   Group "Group" at 455,41 size 373x50
   Button "HmiScreenItemData_8" at 469,45 size 355x40; TextOn 'Back'; TextOff 'Text'
   TextField "Screen title" at 455,41 size 373x50; Text 'Screen title'

screen "BC Max Step Times" 1280x800, template "Template"
   on GenerateScreen: "TitleUpdater"()
   Button "HmiScreenItemData_1" at 1,1 size 150x43; TextOn 'Back'; TextOff 'Commissioning'
      on Release: ActivateScreen("Commissioning Main Page", 0)
   Button "Button_1" at 21,736 size 161x32; TextOff 'Back'
      on Activate: ActivateScreen("IGG Process Times", 0)
   TextField "Text field_25" at 83,285 size 286x22; Text 'Step 040'
   TextField "Text field_29" at 383,118 size 77x20; Text 'Time (ms)'
   TextField "Text field_33" at 83,312 size 286x22; Text 'Step 050'
   IOField "I/O field_58" at 382,312 size 60x22; Authorization "Parameter Change"; FormatPattern s9999999999
      ProcessValue <- "86_Times_STEP_MAX_TIME_STP_050(1)"
   TextField "Text field_35" at 83,367 size 286x22; Text 'Step 070'
   TextField "Text field_65" at 83,144 size 286x22; Text 'Step 001'
   TextField "Text field_67" at 83,173 size 286x22; Text 'Step 005'
   TextField "Text field_69" at 83,200 size 286x22; Text 'Step 010'
   TextField "Text field_71" at 83,229 size 286x22; Text 'Step 020'
   TextField "Text field_73" at 83,257 size 286x22; Text 'Step 030'
   TextField "Text field_42" at 83,118 size 89x20; Text 'Description'
   IOField "I/O field_128" at 382,144 size 60x22; Authorization "Parameter Change"; FormatPattern s9999999999
      ProcessValue <- "86_Times_STEP_MAX_TIME_STP_001(1)"
   IOField "I/O field_133" at 382,173 size 60x22; Authorization "Parameter Change"; FormatPattern s9999999999
      ProcessValue <- "86_Times_STEP_MAX_TIME_STP_005(1)"
   IOField "I/O field_138" at 382,200 size 60x22; Authorization "Parameter Change"; FormatPattern s9999999999
      ProcessValue <- "86_Times_STEP_MAX_TIME_STP_010(1)"
   IOField "I/O field_148" at 382,257 size 60x22; Authorization "Parameter Change"; FormatPattern s9999999999
      ProcessValue <- "86_Times_STEP_MAX_TIME_STP_030(1)"
   IOField "I/O field_64" at 382,367 size 60x22; Authorization "Parameter Change"; FormatPattern s9999999999
      ProcessValue <- "86_Times_STEP_MAX_TIME_STP_070(1)"
   TextField "Text field_53" at 82,92 size 247x26; Text 'BC Maximum Step Times'
   IOField "I/O field_5" at 382,229 size 60x22; Authorization "Parameter Change"; FormatPattern s9999999999
      ProcessValue <- "86_Times_STEP_MAX_TIME_STP_020(1)"
   TextField "Text field_1" at 83,340 size 286x22; Text 'Step 060'
   IOField "I/O field_2" at 382,340 size 60x22; Authorization "Parameter Change"; FormatPattern s9999999999
      ProcessValue <- "86_Times_STEP_MAX_TIME_STP_060(1)"
   TextField "Text field_2" at 461,286 size 286x22; Text 'Step 240'
   TextField "Text field_3" at 750,119 size 77x20; Text 'Time (ms)'
   TextField "Text field_4" at 461,313 size 286x22; Text 'Step 250'
   IOField "I/O field_1" at 758,312 size 60x22; Authorization "Parameter Change"; FormatPattern s9999999999
      ProcessValue <- "86_Times_STEP_MAX_TIME_STP_250(1)"
   TextField "Text field_5" at 461,368 size 286x22; Text 'Step 270'
   TextField "Text field_6" at 461,145 size 286x22; Text 'Step 190'
   TextField "Text field_7" at 461,174 size 286x22; Text 'Step 200'
   TextField "Text field_8" at 461,201 size 286x22; Text 'Step 210'
   TextField "Text field_9" at 461,230 size 286x22; Text 'Step 220'
   TextField "Text field_10" at 461,258 size 286x22; Text 'Step 230'
   TextField "Text field_11" at 461,119 size 89x20; Text 'Description'
   IOField "I/O field_3" at 758,145 size 60x22; Authorization "Parameter Change"; FormatPattern s9999999999
      ProcessValue <- "86_Times_STEP_MAX_TIME_STP_190(1)"
   IOField "I/O field_4" at 758,174 size 60x22; Authorization "Parameter Change"; FormatPattern s9999999999
      ProcessValue <- "86_Times_STEP_MAX_TIME_STP_200(1)"
   IOField "I/O field_6" at 758,201 size 60x22; Authorization "Parameter Change"; FormatPattern s9999999999
      ProcessValue <- "86_Times_STEP_MAX_TIME_STP_210(1)"
   IOField "I/O field_8" at 758,258 size 60x22; Authorization "Parameter Change"; FormatPattern s9999999999
      ProcessValue <- "86_Times_STEP_MAX_TIME_STP_230(1)"
   IOField "I/O field_9" at 758,367 size 60x22; Authorization "Parameter Change"; FormatPattern s9999999999
      ProcessValue <- "86_Times_STEP_MAX_TIME_STP_270(1)"
   IOField "I/O field_10" at 758,230 size 60x22; Authorization "Parameter Change"; FormatPattern s9999999999
      ProcessValue <- "86_Times_STEP_MAX_TIME_STP_220(1)"
   TextField "Text field_13" at 461,341 size 286x22; Text 'Step 260'
   IOField "I/O field_11" at 758,340 size 60x22; Authorization "Parameter Change"; FormatPattern s9999999999
      ProcessValue <- "86_Times_STEP_MAX_TIME_STP_260(1)"
   TextField "Text field_14" at 83,398 size 286x22; Text 'Step 080'
   IOField "I/O field_12" at 382,398 size 60x22; Authorization "Parameter Change"; FormatPattern s9999999999
      ProcessValue <- "86_Times_STEP_MAX_TIME_STP_080(1)"
   TextField "Text field_15" at 83,426 size 286x22; Text 'Step 090'
   IOField "I/O field_13" at 382,426 size 60x22; Authorization "Parameter Change"; FormatPattern s9999999999
      ProcessValue <- "86_Times_STEP_MAX_TIME_STP_090(1)"
   TextField "Text field_16" at 83,453 size 286x22; Text 'Step 100'
   IOField "I/O field_14" at 382,453 size 60x22; Authorization "Parameter Change"; FormatPattern s9999999999
      ProcessValue <- "86_Times_STEP_MAX_TIME_STP_100(1)"
   IOField "I/O field_15" at 382,285 size 60x22; Authorization "Parameter Change"; FormatPattern s9999999999
      ProcessValue <- "86_Times_STEP_MAX_TIME_STP_040(1)"
   TextField "Text field_17" at 461,395 size 286x22; Text 'Step 280'
   IOField "I/O field_16" at 758,394 size 60x22; Authorization "Parameter Change"; FormatPattern s9999999999
      ProcessValue <- "86_Times_STEP_MAX_TIME_STP_280(1)"
   TextField "Text field_18" at 461,426 size 286x22; Text 'Step 290'
   IOField "I/O field_17" at 758,425 size 60x22; Authorization "Parameter Change"; FormatPattern s9999999999
      ProcessValue <- "86_Times_STEP_MAX_TIME_STP_290(1)"
   TextField "Text field_19" at 461,453 size 286x22; Text 'Step 300'
   IOField "I/O field_18" at 758,452 size 60x22; Authorization "Parameter Change"; FormatPattern s9999999999
      ProcessValue <- "86_Times_STEP_MAX_TIME_STP_300(1)"
   TextField "Text field_20" at 461,483 size 286x22; Text 'Step 310'
   IOField "I/O field_19" at 758,482 size 60x22; Authorization "Parameter Change"; FormatPattern s9999999999
      ProcessValue <- "86_Times_STEP_MAX_TIME_STP_310(1)"
   TextField "Text field_21" at 461,510 size 286x22; Text 'Step 320'
   IOField "I/O field_20" at 758,509 size 60x22; Authorization "Parameter Change"; FormatPattern s9999999999
      ProcessValue <- "86_Times_STEP_MAX_TIME_STP_320(1)"
   TextField "Text field_22" at 835,145 size 286x22; Text 'Step 390'
   IOField "I/O field_21" at 1130,144 size 60x22; Authorization "Parameter Change"; FormatPattern s9999999999
      ProcessValue <- "86_Times_STEP_MAX_TIME_STP_390(1)"
   TextField "Text field_23" at 835,118 size 89x20; Text 'Description'
   TextField "Text field_24" at 1122,119 size 77x20; Text 'Time (ms)'
   TextField "Text field_26" at 835,173 size 286x22; Text 'Step 400'
   IOField "I/O field_22" at 1130,172 size 60x22; Authorization "Parameter Change"; FormatPattern s9999999999
      ProcessValue <- "86_Times_STEP_MAX_TIME_STP_400(1)"
   TextField "Text field_27" at 835,200 size 286x22; Text 'Step 410'
   IOField "I/O field_23" at 1130,199 size 60x22; Authorization "Parameter Change"; FormatPattern s9999999999
      ProcessValue <- "86_Times_STEP_MAX_TIME_STP_410(1)"
   TextField "Text field_28" at 835,230 size 286x22; Text 'Step 420'
   IOField "I/O field_24" at 1130,229 size 60x22; Authorization "Parameter Change"; FormatPattern s9999999999
      ProcessValue <- "86_Times_STEP_MAX_TIME_STP_420(1)"
   TextField "Text field_30" at 835,257 size 286x22; Text 'Step 430'
   IOField "I/O field_25" at 1130,256 size 60x22; Authorization "Parameter Change"; FormatPattern s9999999999
      ProcessValue <- "86_Times_STEP_MAX_TIME_STP_430(1)"
   TextField "Text field_31" at 835,285 size 286x22; Text 'Step 440'
   IOField "I/O field_26" at 1130,284 size 60x22; Authorization "Parameter Change"; FormatPattern s9999999999
      ProcessValue <- "86_Times_STEP_MAX_TIME_STP_440(1)"
   TextField "Text field_32" at 835,312 size 286x22; Text 'Step 450'
   IOField "I/O field_27" at 1130,311 size 60x22; Authorization "Parameter Change"; FormatPattern s9999999999
      ProcessValue <- "86_Times_STEP_MAX_TIME_STP_450(1)"
   TextField "Text field_34" at 835,341 size 286x22; Text 'Step 460'
   IOField "I/O field_28" at 1130,340 size 60x22; Authorization "Parameter Change"; FormatPattern s9999999999
      ProcessValue <- "86_Times_STEP_MAX_TIME_STP_460(1)"
   TextField "Text field_36" at 835,369 size 286x22; Text 'Step 470'
   IOField "I/O field_29" at 1130,368 size 60x22; Authorization "Parameter Change"; FormatPattern s9999999999
      ProcessValue <- "86_Times_STEP_MAX_TIME_STP_470(1)"
   TextField "Text field_37" at 835,395 size 286x22; Text 'Step 480'
   IOField "I/O field_30" at 1130,394 size 60x22; Authorization "Parameter Change"; FormatPattern s9999999999
      ProcessValue <- "86_Times_STEP_MAX_TIME_STP_480(1)"
   TextField "Text field_38" at 835,426 size 286x22; Text 'Step 490'
   IOField "I/O field_31" at 1130,425 size 60x22; Authorization "Parameter Change"; FormatPattern s9999999999
      ProcessValue <- "86_Times_STEP_MAX_TIME_STP_490(1)"
   TextField "Text field_39" at 835,452 size 286x22; Text 'Step 500'
   IOField "I/O field_32" at 1130,451 size 60x22; Authorization "Parameter Change"; FormatPattern s9999999999
      ProcessValue <- "86_Times_STEP_MAX_TIME_STP_500(1)"
   TextField "Text field_40" at 835,482 size 286x22; Text 'Step 510'
   IOField "I/O field_33" at 1130,481 size 60x22; Authorization "Parameter Change"; FormatPattern s9999999999
      ProcessValue <- "86_Times_STEP_MAX_TIME_STP_510(1)"
   TextField "Text field_41" at 835,510 size 286x22; Text 'Step 520'
   IOField "I/O field_34" at 1130,509 size 60x22; Authorization "Parameter Change"; FormatPattern s9999999999
      ProcessValue <- "86_Times_STEP_MAX_TIME_STP_520(1)"
   IOField "I/O field_7" at 758,285 size 60x22; Authorization "Parameter Change"; FormatPattern s9999999999
      ProcessValue <- "86_Times_STEP_MAX_TIME_STP_240(1)"
   TextField "Text field_43" at 83,483 size 286x22; Text 'Step 110'
   IOField "I/O field_35" at 382,483 size 60x22; Authorization "Parameter Change"; FormatPattern s9999999999
      ProcessValue <- "86_Times_STEP_MAX_TIME_STP_110(1)"
   TextField "Text field_44" at 83,510 size 286x22; Text 'Step 120'
   IOField "I/O field_36" at 382,510 size 60x22; Authorization "Parameter Change"; FormatPattern s9999999999
      ProcessValue <- "86_Times_STEP_MAX_TIME_STP_120(1)"
   TextField "Text field_45" at 461,538 size 286x22; Text 'Step 330'
   IOField "I/O field_37" at 758,537 size 60x22; Authorization "Parameter Change"; FormatPattern s9999999999
      ProcessValue <- "86_Times_STEP_MAX_TIME_STP_330(1)"
   TextField "Text field_46" at 835,538 size 286x22; Text 'Step 530'
   IOField "I/O field_38" at 1130,537 size 60x22; Authorization "Parameter Change"; FormatPattern s9999999999
      ProcessValue <- "86_Times_STEP_MAX_TIME_STP_530(1)"
   TextField "Text field_47" at 83,538 size 286x22; Text 'Step 130'
   IOField "I/O field_39" at 382,538 size 60x22; Authorization "Parameter Change"; FormatPattern s9999999999
      ProcessValue <- "86_Times_STEP_MAX_TIME_STP_130(1)"
   TextField "Text field_48" at 461,568 size 286x22; Text 'Step 340'
   IOField "I/O field_40" at 758,567 size 60x22; Authorization "Parameter Change"; FormatPattern s9999999999
      ProcessValue <- "86_Times_STEP_MAX_TIME_STP_340(1)"
   TextField "Text field_49" at 835,568 size 286x22; Text 'Step 540'
   IOField "I/O field_41" at 1130,567 size 60x22; Authorization "Parameter Change"; FormatPattern s9999999999
      ProcessValue <- "86_Times_STEP_MAX_TIME_STP_540(1)"
   TextField "Text field_50" at 83,568 size 286x22; Text 'Step 140'
   IOField "I/O field_42" at 382,568 size 60x22; Authorization "Parameter Change"; FormatPattern s9999999999
      ProcessValue <- "86_Times_STEP_MAX_TIME_STP_140(1)"
   TextField "Text field_51" at 461,599 size 286x22; Text 'Step 350'
   IOField "I/O field_43" at 758,598 size 60x22; Authorization "Parameter Change"; FormatPattern s9999999999
      ProcessValue <- "86_Times_STEP_MAX_TIME_STP_350(1)"
   TextField "Text field_52" at 835,599 size 286x22; Text 'Step 550'
   IOField "I/O field_44" at 1130,598 size 60x22; Authorization "Parameter Change"; FormatPattern s9999999999
      ProcessValue <- "86_Times_STEP_MAX_TIME_STP_550(1)"
   TextField "Text field_54" at 83,599 size 286x22; Text 'Step 150'
   IOField "I/O field_45" at 382,599 size 60x22; Authorization "Parameter Change"; FormatPattern s9999999999
      ProcessValue <- "86_Times_STEP_MAX_TIME_STP_150(1)"
   TextField "Text field_55" at 461,628 size 286x22; Text 'Step 360'
   IOField "I/O field_46" at 758,627 size 60x22; Authorization "Parameter Change"; FormatPattern s9999999999
      ProcessValue <- "86_Times_STEP_MAX_TIME_STP_360(1)"
   TextField "Text field_56" at 835,628 size 286x22; Text 'Step 560'
   IOField "I/O field_47" at 1130,627 size 60x22; Authorization "Parameter Change"; FormatPattern s9999999999
      ProcessValue <- "86_Times_STEP_MAX_TIME_STP_560(1)"
   TextField "Text field_57" at 83,628 size 286x22; Text 'Step 160'
   IOField "I/O field_48" at 382,628 size 60x22; Authorization "Parameter Change"; FormatPattern s9999999999
      ProcessValue <- "86_Times_STEP_MAX_TIME_STP_160(1)"
   TextField "Text field_58" at 461,657 size 286x22; Text 'Step 370'
   IOField "I/O field_49" at 758,656 size 60x22; Authorization "Parameter Change"; FormatPattern s9999999999
      ProcessValue <- "86_Times_STEP_MAX_TIME_STP_370(1)"
   TextField "Text field_59" at 835,657 size 286x22; Text 'Step 570'
   IOField "I/O field_50" at 1130,656 size 60x22; Authorization "Parameter Change"; FormatPattern s9999999999
      ProcessValue <- "86_Times_STEP_MAX_TIME_STP_570(1)"
   TextField "Text field_60" at 83,657 size 286x22; Text 'Step 170'
   IOField "I/O field_51" at 382,657 size 60x22; Authorization "Parameter Change"; FormatPattern s9999999999
      ProcessValue <- "86_Times_STEP_MAX_TIME_STP_170(1)"
   TextField "Text field_61" at 461,687 size 286x22; Text 'Step 380'
   IOField "I/O field_52" at 758,686 size 60x22; Authorization "Parameter Change"; FormatPattern s9999999999
      ProcessValue <- "86_Times_STEP_MAX_TIME_STP_380(1)"
   TextField "Text field_63" at 83,687 size 286x22; Text 'Step 180'
   IOField "I/O field_54" at 382,687 size 60x22; Authorization "Parameter Change"; FormatPattern s9999999999
      ProcessValue <- "86_Times_STEP_MAX_TIME_STP_180(1)"
   Group "Group" at 455,41 size 373x50
   Button "HmiScreenItemData_8" at 469,45 size 355x40; TextOn 'Back'; TextOff 'Text'
   TextField "Screen title" at 455,41 size 373x50; Text 'Screen title'

screen "05 Alarm Buffer" 1280x800, template "Template"
   AlarmView "Alarm view_1" at 8,61 size 1258x729
   Button "HmiScreenItemData_2" at 143,2 size 139x43; TextOn 'Back'; TextOff 'Alarm'
      on Release: ActivateScreen("04 Alarm Log", 0)
   Button "HmiScreenItemData_5" at 1,2 size 139x43; TextOn 'Back'; TextOff 'Main Index'
      on Release: ActivateScreen("02 Main Index", 0)
   Button "HmiScreenItemData_4" at 1138,1 size 139x43; TextOn 'I&A Compressor Ok'; TextOff 'Back'
      on Release: function_efd93a16()

screen "08 BTCS MAIN" 1280x800, template "Template"
   Rectangle "Rectangle_1" at 150,160 size 480x40
      Appearance <- "2102_TIME_CALCS_DB_PRE_DWELL_TMR_DN"
   TextField "Text field_4" at 155,165 size 200x30; Text 'Pre-Dwell Time :'
   IOField "I/O field_1" at 360,165 size 60x30; FormatPattern 999
      ProcessValue <- "2110_BTCS_CNTRL_DB_PRE_DWELL_HRS"
   TextField "Text field_5" at 420,165 size 60x30; Text 'Hours'
   IOField "I/O field_2" at 485,165 size 60x30; FormatPattern 99
      ProcessValue <- "2110_BTCS_CNTRL_DB_PRE_DWELL_MINS"
   TextField "Text field_6" at 545,165 size 80x30; Text 'Minutes'
   Rectangle "Rectangle_2" at 150,205 size 480x40
      Appearance <- "2102_TIME_CALCS_DB_DE_OX_TMR_DN"
   TextField "Text field_7" at 155,210 size 200x30; Text 'De-Oxygenate Time :'
   IOField "I/O field_3" at 360,210 size 60x30; FormatPattern 999
      ProcessValue <- "2110_BTCS_CNTRL_DB_DE_OX_HRS"
   TextField "Text field_8" at 420,210 size 60x30; Text 'Hours'
   IOField "I/O field_4" at 485,210 size 60x30; FormatPattern 99
      ProcessValue <- "2110_BTCS_CNTRL_DB_DE_OX_MINS"
   TextField "Text field_9" at 545,210 size 80x30; Text 'Minutes'
   Rectangle "Rectangle_3" at 150,250 size 480x40
      Appearance <- "2102_TIME_CALCS_DB_DWELL_TMR_DN"
   TextField "Text field_10" at 155,255 size 200x30; Text 'Dwell Time :'
   IOField "I/O field_5" at 360,255 size 60x30; FormatPattern 999
      ProcessValue <- "2110_BTCS_CNTRL_DB_DWELL_HRS"
   TextField "Text field_11" at 420,255 size 60x30; Text 'Hours'
   IOField "I/O field_6" at 485,255 size 60x30; FormatPattern 99
      ProcessValue <- "2110_BTCS_CNTRL_DB_DWELL_MINS"
   TextField "Text field_12" at 545,255 size 80x30; Text 'Minutes'
   Rectangle "Rectangle_4" at 150,295 size 480x40
      Appearance <- "2102_TIME_CALCS_DB_RE_OX_TMR_DN"
   TextField "Text field_13" at 155,300 size 200x30; Text 'Re-Oxygenate Time :'
   IOField "I/O field_7" at 360,300 size 60x30; FormatPattern 999
      ProcessValue <- "2110_BTCS_CNTRL_DB_RE_OX_HRS"
   TextField "Text field_14" at 420,300 size 60x30; Text 'Hours'
   IOField "I/O field_8" at 485,300 size 60x30; FormatPattern 99
      ProcessValue <- "2110_BTCS_CNTRL_DB_RE_OX_MINS"
   TextField "Text field_15" at 545,300 size 80x30; Text 'Minutes'
   Rectangle "Rectangle_5" at 150,340 size 480x40
      Appearance <- "2102_TIME_CALCS_DB_POST_DWELL_TMR_DN"
   TextField "Text field_16" at 155,345 size 200x30; Text 'Post-Dwell Time :'
   IOField "I/O field_9" at 360,345 size 60x30; FormatPattern 999
      ProcessValue <- "2110_BTCS_CNTRL_DB_POST_DWELL_HRS"
   TextField "Text field_17" at 420,345 size 60x30; Text 'Hours'
   IOField "I/O field_10" at 485,345 size 60x30; FormatPattern 99
      ProcessValue <- "2110_BTCS_CNTRL_DB_POST_DWELL_MINS"
   TextField "Text field_18" at 545,345 size 80x30; Text 'Minutes'
   Rectangle "Rectangle_6" at 640,205 size 480x40
      Appearance <- "2102_TIME_CALCS_DB_DE_OX_SP_TMR_DN"
   TextField "Text field_19" at 645,210 size 200x30; Text 'At De-Ox Setpoint :'
   IOField "I/O field_11" at 850,210 size 60x30; FormatPattern 999
      ProcessValue <- "2110_BTCS_CNTRL_DB_DE_OX_SP_HRS"
   TextField "Text field_20" at 910,210 size 60x30; Text 'Hours'
   IOField "I/O field_12" at 975,210 size 60x30; FormatPattern 99
      ProcessValue <- "2110_BTCS_CNTRL_DB_DE_OX_SP_MINS"
   TextField "Text field_21" at 1035,210 size 80x30; Text 'Minutes'
   Rectangle "Rectangle_7" at 640,295 size 480x40
      Appearance <- "2102_TIME_CALCS_DB_RE_OX_SP_TMR_DN"
   TextField "Text field_22" at 645,300 size 200x30; Text 'At Re-Ox Setpoint :'
   IOField "I/O field_13" at 850,300 size 60x30; FormatPattern 999
      ProcessValue <- "2110_BTCS_CNTRL_DB_RE_OX_SP_HRS"
   TextField "Text field_23" at 910,300 size 60x30; Text 'Hours'
   IOField "I/O field_14" at 975,300 size 60x30; FormatPattern 99
      ProcessValue <- "2110_BTCS_CNTRL_DB_RE_OX_SP_MINS"
   TextField "Text field_24" at 1035,300 size 80x30; Text 'Minutes'
   TextField "Text field_25" at 155,435 size 200x30; Text 'Total Sequence Time:'
   IOField "I/O field_15" at 360,435 size 60x30; FormatPattern 999
      ProcessValue <- "2110_BTCS_CNTRL_DB_TOT_SEQ_HRS"
   TextField "Text field_26" at 420,435 size 60x30; Text 'Hours'
   IOField "I/O field_16" at 485,435 size 60x30; FormatPattern 99
      ProcessValue <- "2110_BTCS_CNTRL_DB_TOT_SEQ_MINS"
   TextField "Text field_27" at 545,435 size 80x30; Text 'Minutes'
   TextField "Text field_28" at 155,625 size 200x30; Text 'Remaining Time:'
   IOField "I/O field_17" at 360,625 size 60x30; FormatPattern 999
      ProcessValue <- "2110_BTCS_CNTRL_DB_RMNG_SEQ_HRS"
   TextField "Text field_29" at 420,625 size 60x30; Text 'Hours'
   IOField "I/O field_18" at 485,625 size 60x30; FormatPattern 99
      ProcessValue <- "2110_BTCS_CNTRL_DB_RMNG_SEQ_MINS"
   TextField "Text field_30" at 545,625 size 80x30; Text 'Minutes'
   TextField "Text field_61" at 150,575 size 480x35; Text 'INPUT SALINITY'
      Visibility <- "2068_Sys_Status_Data_SAL_VALID"
   TextField "Text field_60" at 150,575 size 480x35; Text 'SALINITY ACCEPTED'
      Visibility <- "2068_Sys_Status_Data_SAL_VALID"
   Button "HmiScreenItemData_1" at 10,10 size 160x50; TextOn 'Back'; TextOff 'Main Index'
      on Release: ActivateScreen("02 Main Index", 0)
   TextField "Text field_1" at 324,55 size 640x35; Text 'BASIC BARGE TWO TANK CONTROL SYSTEM'
   Button "HmiScreenItemData_2" at 1127,4 size 149x50; TextOn 'Back'; TextOff 'Enable'
      on Press: ResetBit("80_From_HMI_RUN_BWTS"); SetBit("80_From_HMI_RUN_BTCS")
      Visibility <- "80_From_HMI_RUN_BTCS"
   Button "HmiScreenItemData_3" at 1127,56 size 149x50; TextOn 'Back'; TextOff 'Disable'
      on Press: ResetBit("80_From_HMI_RUN_BTCS"); SetBit("80_From_HMI_RUN_BWTS")
      Visibility <- "80_From_HMI_RUN_BTCS"
   TextField "Text field_2" at 484,85 size 320x35; Text 'BTCS ENABLED'
      Visibility <- "80_From_HMI_RUN_BTCS"
   TextField "Text field_3" at 484,85 size 320x35; Text 'BTCS DISABLED'
      Visibility <- "80_From_HMI_RUN_BTCS"
   Button "Button_2" at 10,70 size 160x50; TextOn 'User Account'; TextOff 'Alarm Log'; Authorization "User administration"
      on Release: ActivateScreen("04 Alarm Log", 0)
   Group "Group_1" at 150,205 size 480x40
   Group "Group_2" at 150,250 size 480x40
   Group "Group_3" at 150,295 size 480x40
   Group "Group_4" at 150,340 size 480x40
   Group "Group_5" at 640,205 size 480x40
   Group "Group_6" at 640,295 size 480x40
   Group "Group_7" at 150,430 size 480x40
   Group "Group_8" at 150,620 size 480x40
   TextField "Text field_31" at 1005,150 size 120x30; Text 'SETUP'
   TextField "Text field_32" at 1005,420 size 120x30; Text 'CONTROL'
   Button "Button_1" at 150,520 size 230x50; TextOff 'ACCEPT & LAUNCH'
      on Release: ResetBit("2110_BTCS_CNTRL_DB_START_SEQ")
      on Press: SetBit("2110_BTCS_CNTRL_DB_START_SEQ")
      Appearance <- "2110_BTCS_CNTRL_DB_BTCS_STATE"
      Visibility <- "2102_TIME_CALCS_DB_TIMES_VALID"
   SymbolicIOField "Symbolic I/O field_1" at 640,480 size 480x30; TextOn '1'; TextOff '0'; TextList "STATE LIST BTCS"
      ProcessValue <- "2110_BTCS_CNTRL_DB_BTCS_STATE"
   TextField "Text field_33" at 150,480 size 480x35; Text 'TIMES NOT VALID'
      Visibility <- "2102_TIME_CALCS_DB_TIMES_VALID"
   TextField "Text field_34" at 150,480 size 480x35; Text 'TIMES VALID'
      Visibility <- "2102_TIME_CALCS_DB_TIMES_VALID"
   SymbolicIOField "Symbolic I/O field_2" at 640,580 size 480x30; TextOn '1'; TextOff '0'; TextList "STEP LIST BTCS"
      ProcessValue <- "2110_BTCS_CNTRL_DB_BTCS_STEP"
   Button "HmiScreenItemData_4" at 1127,108 size 149x50; TextOn 'Back'; TextOff 'Master Reset'
      on Press: ResetBit("2110_BTCS_CNTRL_DB_RESET_ALL"); SetBit("2110_BTCS_CNTRL_DB_RESET_ALL")
      Visibility <- "80_From_HMI_RUN_BTCS"
   SymbolicIOField "Symbolic I/O field_3" at 360,700 size 140x30; TextOn '1'; TextOff '0'; TextList "Port Tank"
      ProcessValue <- "2110_BTCS_CNTRL_DB_PORT_TANK_STS"
   Button "Button_4" at 150,700 size 180x30; TextOff 'Port Tank'
      on Press: InvertBit("2110_BTCS_CNTRL_DB_PORT_TANK_STS")
      Appearance <- "2110_BTCS_CNTRL_DB_PORT_TANK_STS"
   TextField "Text field_35" at 1025,690 size 100x30; Text 'TANKS'
   SymbolicIOField "Symbolic I/O field_4" at 360,740 size 140x30; TextOn '1'; TextOff '0'; TextList "Port Tank"
      ProcessValue <- "2110_BTCS_CNTRL_DB_STBD_TANK_STS"
   Button "Button_5" at 150,740 size 180x30; TextOff 'Starboard Tank'
      on Press: InvertBit("2110_BTCS_CNTRL_DB_STBD_TANK_STS")
      Appearance <- "2110_BTCS_CNTRL_DB_STBD_TANK_STS"
   TextField "Text field_37" at 515,700 size 60x30; Text 'O2 :'
   IOField "I/O field_20" at 575,700 size 60x30; FormatPattern 99.99
      ProcessValue <- "20_TANKS_IP_DATA_RIO_02_FIRST_TANK_BWT_DO"
   TextField "Text field_36" at 640,700 size 60x30; Text 'ph :'
   IOField "I/O field_19" at 700,700 size 60x30; FormatPattern 99.99
      ProcessValue <- "20_TANKS_IP_DATA_RIO_02_FIRST_TANK_BWT_PH"
   TextField "Text field_38" at 775,700 size 65x30; Text 'Temp :'
   IOField "I/O field_21" at 840,700 size 60x30; FormatPattern 99.99
      ProcessValue <- "20_TANKS_IP_DATA_RIO_02_FIRST_TANK_BWT_TEMP"
   TextField "Text field_39" at 910,700 size 65x30; Text 'Level :'
   IOField "I/O field_22" at 975,700 size 60x30; FormatPattern 99.9
      ProcessValue <- "20_TANKS_IP_DATA_RIO_02_FIRST_TANK_BWT_LEVEL"
   TextField "Text field_40" at 515,740 size 60x30; Text 'O2 :'
   IOField "I/O field_23" at 575,740 size 60x30; FormatPattern 99.99
      ProcessValue <- "20_TANKS_IP_DATA_RIO_02_SECOND_TANK_BWT_DO"
   TextField "Text field_41" at 640,740 size 60x30; Text 'ph :'
   IOField "I/O field_24" at 700,740 size 60x30; FormatPattern 99.99
      ProcessValue <- "20_TANKS_IP_DATA_RIO_02_SECOND_TANK_BWT_PH"
   TextField "Text field_42" at 775,740 size 65x30; Text 'Temp :'
   IOField "I/O field_25" at 840,740 size 60x30; FormatPattern 99.99
      ProcessValue <- "20_TANKS_IP_DATA_RIO_02_SECOND_TANK_BWT_TEMP"
   TextField "Text field_43" at 910,740 size 65x30; Text 'Level :'
   IOField "I/O field_26" at 975,740 size 60x30; FormatPattern 99.9
      ProcessValue <- "20_TANKS_IP_DATA_RIO_02_SECOND_TANK_BWT_LEVEL"
   Group "Group" at 150,160 size 480x40
   Group "Group_9" at 150,160 size 480x40
   Group "Group_10" at 150,340 size 480x40
   Group "Group_12" at 150,295 size 480x40
   Group "Group_13" at 640,205 size 480x40
   Group "Group_14" at 150,250 size 480x40
   Group "Group_15" at 150,205 size 480x40
   Group "Group_16" at 640,295 size 480x40
   Rectangle "Rectangle_15" at 249,485 size 303x130
      Visibility <- "2100_AUTO_SEQ_DB_SEQ_RNG"
   Button "Button_3" at 400,520 size 230x50; TextOff 'ABORT - STOP'
      on Release: ResetBit("2110_BTCS_CNTRL_DB_STOP_SEQ")
      on Press: SetBit("2110_BTCS_CNTRL_DB_STOP_SEQ")
      Appearance <- "2110_BTCS_CNTRL_DB_BTCS_STATE"
   Group "Group_17" at 640,250 size 480x40
   Group "Group_18" at 640,250 size 480x40
   Group "Group_11" at 647,276 size 480x40
   Group "Group_19" at 1083,420 size 47x365
   Rectangle "Rectangle_13" at 150,160 size 480x40
      Appearance <- "2102_TIME_CALCS_DB_PRE_DWELL_TMR_DN"
      Visibility <- "2100_AUTO_SEQ_DB_SEQ_RNG"
   TextField "Text field_44" at 155,165 size 310x30; Text 'Pre-Dwell Time Remaining :'
      Visibility <- "2100_AUTO_SEQ_DB_SEQ_RNG"
   IOField "I/O field_28" at 465,165 size 80x30; FormatPattern 999999
      ProcessValue <- "2102_TIME_CALCS_DB_PRE_DWELL_MINS_RMNG"
      Visibility <- "2100_AUTO_SEQ_DB_SEQ_RNG"
   TextField "Text field_46" at 545,165 size 80x30; Text 'Minutes'
      Visibility <- "2100_AUTO_SEQ_DB_SEQ_RNG"
   Rectangle "Rectangle_14" at 150,340 size 480x40
      Visibility <- "2100_AUTO_SEQ_DB_SEQ_RNG"
      Appearance <- "2102_TIME_CALCS_DB_POST_DWELL_TMR_DN"
   TextField "Text field_45" at 155,345 size 310x30; Text 'Post-Dwell Time Remaining :'
      Visibility <- "2100_AUTO_SEQ_DB_SEQ_RNG"
   IOField "I/O field_27" at 465,345 size 80x30; FormatPattern 999999
      Visibility <- "2100_AUTO_SEQ_DB_SEQ_RNG"
      ProcessValue <- "2102_TIME_CALCS_DB_POST_DWELL_MINS_RMNG"
   TextField "Text field_47" at 545,345 size 80x30; Text 'Minutes'
      Visibility <- "2100_AUTO_SEQ_DB_SEQ_RNG"
   Rectangle "Rectangle_16" at 150,295 size 480x40
      Visibility <- "2100_AUTO_SEQ_DB_SEQ_RNG"
      Appearance <- "2102_TIME_CALCS_DB_RE_OX_TMR_DN"
   TextField "Text field_50" at 155,300 size 310x30; Text 'Re-Oxygenate Time Remaining :'
      Visibility <- "2100_AUTO_SEQ_DB_SEQ_RNG"
   IOField "I/O field_30" at 465,300 size 80x30; FormatPattern 999999
      Visibility <- "2100_AUTO_SEQ_DB_SEQ_RNG"
      ProcessValue <- "2102_TIME_CALCS_DB_RE_OX_MINS_RMNG"
   TextField "Text field_51" at 545,300 size 80x30; Text 'Minutes'
      Visibility <- "2100_AUTO_SEQ_DB_SEQ_RNG"
   Rectangle "Rectangle_17" at 640,205 size 480x40
      Visibility <- "2100_AUTO_SEQ_DB_SEQ_RNG"
      Appearance <- "2102_TIME_CALCS_DB_DE_OX_SP_TMR_DN"
   TextField "Text field_52" at 645,210 size 310x30; Text 'At De-Ox Time Remaining :'
      Visibility <- "2100_AUTO_SEQ_DB_SEQ_RNG"
   IOField "I/O field_31" at 955,210 size 80x30; FormatPattern 999999
      Visibility <- "2100_AUTO_SEQ_DB_SEQ_RNG"
      ProcessValue <- "2102_TIME_CALCS_DB_DE_OX_SP_MINS_RMNG"
   TextField "Text field_53" at 1035,210 size 80x30; Text 'Minutes'
      Visibility <- "2100_AUTO_SEQ_DB_SEQ_RNG"
   Rectangle "Rectangle_18" at 150,250 size 480x40
      Visibility <- "2100_AUTO_SEQ_DB_SEQ_RNG"
      Appearance <- "2102_TIME_CALCS_DB_DWELL_TMR_DN"
   TextField "Text field_54" at 155,255 size 310x30; Text 'Dwell Time Remaining :'
      Visibility <- "2100_AUTO_SEQ_DB_SEQ_RNG"
   IOField "I/O field_32" at 465,255 size 80x30; FormatPattern 999999
      Visibility <- "2100_AUTO_SEQ_DB_SEQ_RNG"
      ProcessValue <- "2102_TIME_CALCS_DB_DWELL_MINS_RMNG"
   TextField "Text field_55" at 545,255 size 80x30; Text 'Minutes'
      Visibility <- "2100_AUTO_SEQ_DB_SEQ_RNG"
   Rectangle "Rectangle_19" at 150,205 size 480x40
      Visibility <- "2100_AUTO_SEQ_DB_SEQ_RNG"
      Appearance <- "2102_TIME_CALCS_DB_DE_OX_TMR_DN"
   TextField "Text field_56" at 155,210 size 310x30; Text 'De-Oxygenate Time Remaining :'
      Visibility <- "2100_AUTO_SEQ_DB_SEQ_RNG"
   IOField "I/O field_33" at 465,210 size 80x30; FormatPattern 999999
      Visibility <- "2100_AUTO_SEQ_DB_SEQ_RNG"
      ProcessValue <- "2102_TIME_CALCS_DB_DE_OX_MINS_RMNG"
   TextField "Text field_57" at 545,210 size 80x30; Text 'Minutes'
      Visibility <- "2100_AUTO_SEQ_DB_SEQ_RNG"
   Rectangle "Rectangle_20" at 640,295 size 480x40
      Visibility <- "2100_AUTO_SEQ_DB_SEQ_RNG"
      Appearance <- "2102_TIME_CALCS_DB_RE_OX_SP_TMR_DN"
   TextField "Text field_58" at 645,300 size 310x30; Text 'At Re-Ox Time Remaining :'
      Visibility <- "2100_AUTO_SEQ_DB_SEQ_RNG"
   IOField "I/O field_34" at 955,300 size 80x30; FormatPattern 999999
      Visibility <- "2100_AUTO_SEQ_DB_SEQ_RNG"
      ProcessValue <- "2102_TIME_CALCS_DB_RE_OX_SP_MINS_RMNG"
   TextField "Text field_59" at 1035,300 size 80x30; Text 'Minutes'
      Visibility <- "2100_AUTO_SEQ_DB_SEQ_RNG"
   Rectangle "Rectangle_21" at 640,250 size 480x40
      Appearance <- "2068_Sys_Status_Data_SAL_VALID"
   TextField "Text field_48" at 645,255 size 200x30; Text 'Set Salinity Value :'
   IOField "I/O field_29" at 850,255 size 90x30; FormatPattern 99.9; Unit psu
      ProcessValue <- "80_From_HMI_SAL_VALUE"
   Button "HmiScreenItemData_5" at 955,255 size 150x30; TextOn 'Back'; TextOff 'Confirm Salinity'
      on Press: function_b14e0dd5("80_From_HMI_SAL_CNFRM", 0)
   Rectangle "Rectangle_22" at 647,276 size 480x40
      Visibility <- "2100_AUTO_SEQ_DB_SEQ_RNG"
      Appearance <- "2102_TIME_CALCS_DB_RE_OX_SP_TMR_DN"
   TextField "Text field_49" at 652,281 size 310x30; Text 'Salinity Value :'
      Visibility <- "2100_AUTO_SEQ_DB_SEQ_RNG"
   IOField "I/O field_36" at 962,281 size 90x30; FormatPattern 99.9; Unit psu
      ProcessValue <- "80_From_HMI_SAL_VALUE"
      Visibility <- "2100_AUTO_SEQ_DB_SEQ_RNG"
   Rectangle "Rectangle_23" at 640,250 size 480x40
      Visibility <- "2068_Sys_Status_Data_SAL_CNF_CHK"
   TextField "Text field_62" at 645,255 size 250x30; Text 'Salinity Value < 1 Confirm? :'
      Visibility <- "2068_Sys_Status_Data_SAL_CNF_CHK"
   Button "Button_6" at 910,255 size 80x30; TextOff 'YES'
      Visibility <- "2068_Sys_Status_Data_SAL_CNF_CHK"
      on Press: function_b14e0dd5("80_From_HMI_LOW_SAL_ACPT", 0)
   Button "Button_7" at 1020,255 size 80x30; TextOff 'NO'
      Visibility <- "2068_Sys_Status_Data_SAL_CNF_CHK"
      on Press: function_b14e0dd5("80_From_HMI_LOW_SAL_RJCT", 0)
   Rectangle "Rectangle_24" at 1083,420 size 47x365
      Visibility <- "2068_Sys_Status_Data_SAL_CNF_CHK"
   TextField "Text field_65" at 1084,450 size 46x80; Text '!!! WARNING Salinity < 1 Outside Of Certified Range !!!'
      Visibility <- "2068_Sys_Status_Data_SAL_CNF_CHK"
   TextField "Text field_66" at 1084,550 size 46x80; Text 'Confirming Above Means :'
      Visibility <- "2068_Sys_Status_Data_SAL_CNF_CHK"
   TextField "Text field_67" at 1084,650 size 46x80; Text '!!! User Takes Responsability For This Action !!!'
      Visibility <- "2068_Sys_Status_Data_SAL_CNF_CHK"

screen "BC Digital Inputs" 1280x800, template "Template"
   on GenerateScreen: "TitleUpdater"()
   Button "HmiScreenItemData_1" at 1,1 size 150x43; TextOn 'Back'; TextOff 'Commissioning'
      on Release: ActivateScreen("Commissioning Main Page", 0)
   TextField "Text field_37" at 361,69 size 287x26; Text 'Burner Control PLC (Rack 2)'
   TextField "Text field_38" at 361,139 size 55x22; Text 'I0.0'
   TextField "Text field_39" at 361,174 size 55x22; Text 'I0.1'
   TextField "Text field_40" at 361,210 size 55x22; Text 'I0.2'
   TextField "Text field_41" at 361,246 size 55x22; Text 'I0.3'
   TextField "Text field_42" at 361,282 size 55x22; Text 'I0.4'
   TextField "Text field_43" at 361,318 size 55x22; Text 'I0.5'
   TextField "Text field_44" at 361,354 size 55x22; Text 'I0.6'
   TextField "Text field_45" at 361,390 size 55x22; Text 'I0.7'
   Circle "Circle_33" at 421,139 size 20x20
      Appearance <- "10 DI_DATA_PS101"
   Circle "Circle_34" at 421,175 size 20x20
      Appearance <- "10 DI_DATA_E131_SHTDN"
   Circle "Circle_35" at 421,211 size 20x20
      Appearance <- "10 DI_DATA_R2_SPR_DI_0_2"
   Circle "Circle_36" at 421,247 size 20x20
      Appearance <- "10 DI_DATA_R2_SPR_DI_0_3"
   Circle "Circle_37" at 421,282 size 20x20
      Appearance <- "10 DI_DATA_X001_PWR_OK"
   Circle "Circle_38" at 421,318 size 20x20
      Appearance <- "10 DI_DATA_FD001_PWR_OK"
   Circle "Circle_39" at 421,354 size 20x20
      Appearance <- "10 DI_DATA_FD001_OK"
   Circle "Circle_40" at 421,390 size 20x20
      Appearance <- "103_Main_Burner_DB_DN_OK(1)"
   TextField "Text field_46" at 378,107 size 49x26; Text 'I0'
   TextField "Text field_47" at 361,458 size 55x22; Text 'I1.0'
   TextField "Text field_48" at 361,493 size 55x22; Text 'I1.1'
   TextField "Text field_49" at 361,529 size 55x22; Text 'I1.2'
   TextField "Text field_50" at 361,565 size 55x22; Text 'I1.3'
   TextField "Text field_51" at 361,601 size 55x22; Text 'I1.4'
   TextField "Text field_52" at 361,637 size 55x22; Text 'I1.5'
   TextField "Text field_53" at 361,673 size 55x22; Text 'I1.6'
   TextField "Text field_54" at 361,709 size 55x22; Text 'I1.7'
   Circle "Circle_41" at 421,458 size 20x20
      Appearance <- "10 DI_DATA_FS123"
   Circle "Circle_42" at 421,494 size 20x20
      Appearance <- "10 DI_DATA_FS115(1)"
   Circle "Circle_43" at 421,530 size 20x20
      Appearance <- "10 DI_DATA_FS320"
   Circle "Circle_44" at 421,566 size 20x20
      Appearance <- "10 DI_DATA_FS317"
   Circle "Circle_45" at 421,601 size 20x20
      Appearance <- "10 DI_DATA_P301_TRIPPED(1)"
   Circle "Circle_46" at 421,637 size 20x20
      Appearance <- "10 DI_DATA_P301_ENBLD"
   Circle "Circle_47" at 421,673 size 20x20
      Appearance <- "10 DI_DATA_R2_SPR_DI_1_6"
   Circle "Circle_48" at 421,709 size 20x20
      Appearance <- "10 DI_DATA_ESD_OK"
   TextField "Text field_55" at 378,426 size 49x26; Text 'I1'
   TextField "Text field_56" at 652,139 size 55x22; Text 'I2.0'
   TextField "Text field_57" at 652,174 size 55x22; Text 'I2.1'
   TextField "Text field_58" at 652,210 size 55x22; Text 'I2.2'
   TextField "Text field_59" at 652,246 size 55x22; Text 'I2.3'
   TextField "Text field_60" at 652,282 size 55x22; Text 'I2.4'
   TextField "Text field_61" at 652,318 size 55x22; Text 'I2.5'
   TextField "Text field_62" at 652,354 size 55x22; Text 'I2.6'
   TextField "Text field_63" at 652,390 size 55x22; Text 'I2.7'
   Circle "Circle_49" at 712,139 size 20x20
      Appearance <- "10 DI_DATA_E600_NOK"
   Circle "Circle_50" at 712,175 size 20x20
      Appearance <- "10 DI_DATA_E600_HIHI"
   Circle "Circle_51" at 712,211 size 20x20
      Appearance <- "10 DI_DATA_E600_LOLO"
   Circle "Circle_52" at 712,247 size 20x20
      Appearance <- "10 DI_DATA_E600_PWR_OK"
   Circle "Circle_53" at 712,282 size 20x20
      Appearance <- "10 DI_DATA_E700_PWR_OK"
   Circle "Circle_54" at 712,318 size 20x20
      Appearance <- "10 DI_DATA_E700_OPACITY"
   Circle "Circle_55" at 712,354 size 20x20
      Appearance <- "10 DI_DATA_TS403_FAULT(1)"
   Circle "Circle_56" at 712,390 size 20x20
      Appearance <- "10 DI_DATA_TS006"
   TextField "Text field_64" at 669,107 size 49x26; Text 'I2'
   TextField "Text field_65" at 650,458 size 55x22; Text 'I3.0'
   TextField "Text field_66" at 650,493 size 55x22; Text 'I3.1'
   TextField "Text field_67" at 650,529 size 55x22; Text 'I3.2'
   TextField "Text field_68" at 650,565 size 55x22; Text 'I3.3'
   TextField "Text field_69" at 650,601 size 55x22; Text 'I3.4'
   TextField "Text field_70" at 650,637 size 55x22; Text 'I3.5'
   TextField "Text field_71" at 650,673 size 55x22; Text 'I3.6'
   TextField "Text field_72" at 650,709 size 55x22; Text 'I3.7'
   Circle "Circle_57" at 710,458 size 20x20
      Appearance <- "10 DI_DATA_S2_8K1_OK"
   Circle "Circle_58" at 710,494 size 20x20
      Appearance <- "10 DI_DATA_E131_WRNG"
   Circle "Circle_59" at 710,530 size 20x20
      Appearance <- "10 DI_DATA_R2_SPR_DI_3_2"
   Circle "Circle_60" at 710,566 size 20x20
      Appearance <- "10 DI_DATA_E131_OK"
   Circle "Circle_61" at 710,601 size 20x20
      Appearance <- "10 DI_DATA_LS001"
   Circle "Circle_62" at 710,637 size 20x20
      Appearance <- "10 DI_DATA_P305_TRIPPED"
   Circle "Circle_63" at 710,673 size 20x20
      Appearance <- "10 DI_DATA_P305_ENBLD"
   Circle "Circle_64" at 710,709 size 20x20
      Appearance <- "10 DI_DATA_R2_SPR_DI_3_7"
   TextField "Text field_73" at 667,426 size 49x26; Text 'I3'
   TextField "Text field_107" at 450,138 size 180x22; Text 'CA Pressure Switch PS101'
   TextField "Text field_108" at 450,176 size 180x22; Text 'IA Comp Shutdown E131'
   TextField "Text field_109" at 449,216 size 180x22; Text 'Spare Input'
   TextField "Text field_110" at 449,250 size 180x22; Text 'Spare Input'
   TextField "Text field_111" at 449,282 size 180x22; Text 'Ignitor Power Healthy X001'
   TextField "Text field_112" at 449,317 size 180x22; Text 'FDU Power Healthy FD001'
   TextField "Text field_113" at 449,353 size 180x22; Text 'FDU Healthy FD001'
   TextField "Text field_114" at 449,390 size 180x22; Text 'Burner Flame Detected FD001'
   TextField "Text field_116" at 447,458 size 180x22; Text 'Pilot Ign. Air Flow Sw FS123'
   TextField "Text field_117" at 447,494 size 180x22; Text 'Main Atom Air Flow Sw FS115'
   TextField "Text field_118" at 447,529 size 180x22; Text 'Nozzle CW Flow Sw FS320'
   TextField "Text field_119" at 447,566 size 180x22; Text 'Jacket CW Flow Sw FS317'
   TextField "Text field_120" at 447,602 size 180x22; Text 'CSW Pump Tripped P301'
   TextField "Text field_121" at 447,637 size 180x22; Text 'CSW Pump Enabled P301'
   TextField "Text field_122" at 447,710 size 180x22; Text 'Ext. Shutdown'
   TextField "Text field_123" at 740,137 size 180x22; Text 'O2 System Fail E600'
   TextField "Text field_124" at 740,174 size 180x22; Text 'O2 Hi Hi E600'
   TextField "Text field_125" at 739,210 size 180x22; Text 'O2 Lo Lo E600'
   TextField "Text field_126" at 739,246 size 180x22; Text 'O2 System Power Healthy E600'
   TextField "Text field_127" at 739,280 size 180x22; Text 'Soot System Power Healthy E700'
   TextField "Text field_128" at 739,315 size 180x22; Text 'Soot System Opacity E700'
   TextField "Text field_129" at 739,352 size 180x22; Text 'IG Temp Hi Hi Switch TS403'
   TextField "Text field_130" at 740,390 size 180x22; Text 'IG Shell Temp Hi Switch TS006'
   TextField "Text field_131" at 739,458 size 180x22; Text 'IGG E-Stop Healthy'
   TextField "Text field_132" at 739,493 size 180x22; Text 'IA Comp Warning E131'
   TextField "Text field_133" at 739,529 size 180x22; Text 'Spare Input'
   TextField "Text field_134" at 739,637 size 180x22; Text 'Fresh Water Pump Tripped P305'
   TextField "Text field_135" at 739,673 size 180x22; Text 'Fresh Water Pump Enabled P305'
   TextField "Text field_136" at 739,709 size 180x22; Text 'Spare Input'
   TextField "Text field_137" at 739,565 size 180x22; Text 'IA Comp Healthy E131'
   TextField "Text field_138" at 739,601 size 180x22; Text 'Shell CW Level Hi Hi Sw LS001'
   TextField "Text field_115" at 447,673 size 180x22; Text 'Spare Input'
   Group "Group" at 740,44 size 373x50
   Button "HmiScreenItemData_8" at 754,48 size 355x40; TextOn 'Back'; TextOff 'Text'
   TextField "Screen title" at 740,44 size 373x50; Text 'Screen title'

screen "GCU Digital Inputs" 1280x800, template "Template"
   on GenerateScreen: "TitleUpdater"()
   Button "HmiScreenItemData_1" at 1,1 size 150x43; TextOn 'Back'; TextOff 'Commissioning'
      on Release: ActivateScreen("Commissioning Main Page", 0)
   AlarmView "Alarm view_1" at 0,777 size 1280x23
   TextField "Text field_37" at 165,44 size 300x30; Text 'GCU Control PLC (Rack 3)'
   TextField "Text field_34" at 745,74 size 60x30; Text 'I 2'
   TextField "Text field_35" at 745,384 size 70x22; Text 'I 138.7'
   Circle "Circle_16" at 825,384 size 20x20
      Appearance <- "10_DI_DATA_P_303_ENBLD"
   TextField "Text field_36" at 865,384 size 230x22; Text 'P303 ENABLED'
   TextField "Text field_39" at 745,344 size 70x22; Text 'I 138.6'
   Circle "Circle_17" at 825,344 size 20x20
      Appearance <- "10_DI_DATA_EPB_8S1"
   TextField "Text field_40" at 865,344 size 230x22; Text 'PB E-STOP'
   TextField "Text field_41" at 745,304 size 70x22; Text 'I 138.5'
   Circle "Circle_18" at 825,304 size 20x20
      Appearance <- "10_DI_DATA_PB_10S2"
   TextField "Text field_42" at 865,304 size 230x22; Text 'PB STOP'
   TextField "Text field_43" at 745,264 size 70x22; Text 'I 138.4'
   Circle "Circle_19" at 825,264 size 20x20
      Appearance <- "10_DI_DATA_PB_10S1"
   TextField "Text field_44" at 865,264 size 230x22; Text 'PB START'
   TextField "Text field_45" at 745,224 size 70x22; Text 'I 138.3'
   Circle "Circle_20" at 825,224 size 20x20
      Appearance <- "10_DI_DATA_P_304_ENBLD"
   TextField "Text field_46" at 865,224 size 230x22; Text 'P304 ENABLED'
   TextField "Text field_47" at 745,184 size 70x22; Text 'I 138.2'
   Circle "Circle_21" at 825,184 size 20x20
      Appearance <- "10_DI_DATA_LS_303_LO"
   TextField "Text field_48" at 863,184 size 230x22; Text 'LS303 GCU LOW LEVEL'
   TextField "Text field_49" at 745,144 size 70x22; Text 'I 138.1'
   Circle "Circle_22" at 825,144 size 20x20
      Appearance <- "10_DI_DATA_CV441_CLSD"
   TextField "Text field_50" at 865,144 size 230x22; Text 'CV441 CLOSED'
   TextField "Text field_51" at 745,104 size 70x22; Text 'I 138.0'
   Circle "Circle_23" at 825,104 size 20x20
      Appearance <- "10_DI_DATA_CV441_OPN"
   TextField "Text field_52" at 865,104 size 230x22; Text 'CV441 OPEN'
   TextField "Text field_53" at 745,424 size 60x30; Text 'I 3'
   TextField "Text field_54" at 745,734 size 70x22; Text 'I 139.7'
   Circle "Circle_24" at 825,734 size 20x20
      Appearance <- "10_DI_DATA_E_400_NOK"
   TextField "Text field_55" at 865,734 size 230x22; Text 'E400 FAULT'
   TextField "Text field_56" at 745,694 size 70x22; Text 'I 139.6'
   Circle "Circle_25" at 825,694 size 20x20
      Appearance <- "10_DI_DATA_E_400_RUN"
   TextField "Text field_57" at 865,694 size 230x22; Text 'E400 LOADED'
   TextField "Text field_58" at 745,654 size 70x22; Text 'I 139.5'
   Circle "Circle_26" at 825,654 size 20x20
      Appearance <- "10_DI_DATA_P_304_OK"
   TextField "Text field_59" at 865,654 size 230x22; Text 'P304 HEALTHY'
   TextField "Text field_60" at 745,614 size 70x22; Text 'I 139.4'
   Circle "Circle_27" at 825,614 size 20x20
      Appearance <- "10_DI_DATA_6Q6_PWR_OK"
   TextField "Text field_61" at 865,614 size 230x22; Text 'PANEL VENT POWER OK'
   TextField "Text field_62" at 745,574 size 70x22; Text 'I 139.3'
   Circle "Circle_28" at 825,574 size 20x20
      Appearance <- "10_DI_DATA_5T1_PWR_OK"
   TextField "Text field_63" at 865,574 size 230x22; Text '5T1 POWER OK'
   TextField "Text field_64" at 745,534 size 70x22; Text 'I 139.2'
   Circle "Circle_29" at 825,534 size 20x20
      Appearance <- "10_DI_DATA_P_303_OK"
   TextField "Text field_65" at 865,534 size 230x22; Text 'P303 HEALTHY'
   TextField "Text field_66" at 745,494 size 70x22; Text 'I 139.1'
   Circle "Circle_30" at 825,494 size 20x20
      Appearance <- "10_DI_DATA_E_400_SHTDN"
   TextField "Text field_67" at 865,494 size 230x22; Text 'E400 TRIPPED / FAULT'
   TextField "Text field_68" at 745,454 size 70x22; Text 'I 139.0'
   Circle "Circle_31" at 825,454 size 20x20
      Appearance <- "Process Gas Compressor Running/Stopped"
   TextField "Text field_69" at 865,454 size 230x22; Text 'E400 RUN / STOP'
   TextField "Text field_1" at 165,74 size 60x30; Text 'I 0'
   TextField "Text field_15" at 165,384 size 70x22; Text 'I 136.7'
   Circle "Circle_7" at 245,384 size 20x20
      Appearance <- "10_DI_DATA_CV341_CLSD"
   TextField "Text field_16" at 285,384 size 230x22; Text 'CV341 CLOSED'
   TextField "Text field_13" at 165,344 size 70x22; Text 'I 136.6'
   Circle "Circle_6" at 245,344 size 20x20
      Appearance <- "10_DI_DATA_CV341_OPN"
   TextField "Text field_14" at 285,344 size 230x22; Text 'CV341 OPEN'
   TextField "Text field_11" at 165,304 size 70x22; Text 'I 136.5'
   Circle "Circle_5" at 245,304 size 20x20
      Appearance <- "10_DI_DATA_FS_350_FLW_OK"
   TextField "Text field_12" at 285,304 size 230x22; Text 'FS350 FCW FLOW'
   TextField "Text field_9" at 165,264 size 70x22; Text 'I 136.4'
   Circle "Circle_4" at 245,264 size 20x20
      Appearance <- "10_DI_DATA_CV358_CLSD"
   TextField "Text field_10" at 285,264 size 230x22; Text 'CV358 CLOSED'
   TextField "Text field_7" at 165,224 size 70x22; Text 'I 136.3'
   Circle "Circle_3" at 245,224 size 20x20
      Appearance <- "10_DI_DATA_CV358_OPN"
   TextField "Text field_8" at 285,224 size 230x22; Text 'CV358 OPEN'
   TextField "Text field_5" at 165,184 size 70x22; Text 'I 136.2'
   Circle "Circle_2" at 245,184 size 20x20
      Appearance <- "10_DI_DATA_FS_332 FLW_OK"
   TextField "Text field_6" at 285,184 size 230x22; Text 'FS332 CSW FLOW'
   TextField "Text field_3" at 165,144 size 70x22; Text 'I 136.1'
   Circle "Circle_1" at 245,144 size 20x20
      Appearance <- "10_DI_DATA_R3_SPR_DI_136_1"
   TextField "Text field_4" at 285,144 size 230x22; Text 'R3_SPR_DI_136_1'
   TextField "Text field_38" at 165,104 size 70x22; Text 'I 136.0'
   Circle "Circle_33" at 245,104 size 20x20
      Appearance <- "10_DI_DATA_R3_SPR_DI_136_0"
   TextField "Text field_2" at 285,104 size 230x22; Text 'R3_SPR_DI_136_0'
   TextField "Text field_17" at 165,424 size 60x30; Text 'I 1'
   TextField "Text field_18" at 165,734 size 70x22; Text 'I 137.7'
   Circle "Circle_8" at 245,734 size 20x20
      Appearance <- "10_DI_DATA_CV409_CLSD"
   TextField "Text field_19" at 285,734 size 230x22; Text 'CV409 CLOSED'
   TextField "Text field_20" at 165,694 size 70x22; Text 'I 137.6'
   Circle "Circle_9" at 245,694 size 20x20
      Appearance <- "10_DI_DATA_CV409_OPN"
   TextField "Text field_21" at 285,694 size 230x22; Text 'CV409 OPEN'
   TextField "Text field_22" at 165,654 size 70x22; Text 'I 137.5'
   Circle "Circle_10" at 245,654 size 20x20
      Appearance <- "10_DI_DATA_CV411_CLSD"
   TextField "Text field_23" at 285,654 size 230x22; Text 'CV411 CLOSED'
   TextField "Text field_24" at 165,614 size 70x22; Text 'I 137.4'
   Circle "Circle_11" at 245,614 size 20x20
      Appearance <- "10_DI_DATA_CV411_OPN"
   TextField "Text field_25" at 285,614 size 230x22; Text 'CV411 OPEN'
   TextField "Text field_26" at 165,574 size 70x22; Text 'I 137.3'
   Circle "Circle_12" at 245,574 size 20x20
      Appearance <- "10_DI_DATA_CV407_CLSD"
   TextField "Text field_27" at 285,574 size 230x22; Text 'CV407 CLOSED'
   TextField "Text field_28" at 165,534 size 70x22; Text 'I 137.2'
   Circle "Circle_13" at 245,534 size 20x20
      Appearance <- "10_DI_DATA_CV407_OPN"
   TextField "Text field_29" at 285,534 size 230x22; Text 'CV407 OPEN'
   TextField "Text field_30" at 165,494 size 70x22; Text 'I 137.1'
   Circle "Circle_14" at 245,494 size 20x20
      Appearance <- "10_DI_DATA_CV406_CLSD"
   TextField "Text field_31" at 285,494 size 230x22; Text 'CV406 CLOSED'
   TextField "Text field_32" at 165,454 size 70x22; Text 'I 137.0'
   Circle "Circle_15" at 245,454 size 20x20
      Appearance <- "10_DI_DATA_CV406_OPN"
   TextField "Text field_33" at 285,454 size 230x22; Text 'CV406 OPEN'
   Group "Group_1" at 851,41 size 373x50
   Button "HmiScreenItemData_8" at 865,45 size 355x40; TextOn 'Back'; TextOff 'Text'
   TextField "Screen title" at 851,41 size 373x50; Text 'Screen title'

